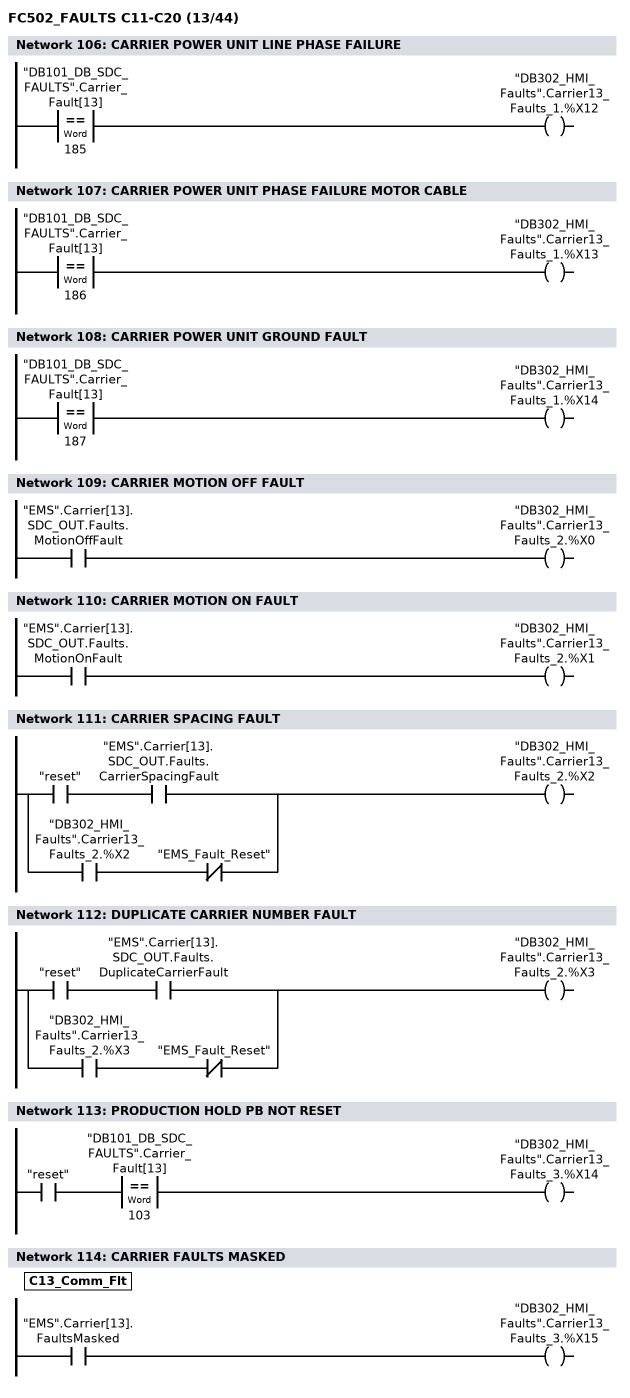
   RUNG wire#powerrail
      { S7_Templates := "SrcType := Word" } EQ_Contact(in1 := "DB101_DB_SDC_FAULTS".Carrier_Fault[13], in2 := 185)
      Coil( "DB302_HMI_Faults".Carrier13_Faults_1.%X12 )
   END_RUNG
   // the same network as SCL:
   "DB302_HMI_Faults".Carrier13_Faults_1.%X12 := "DB101_DB_SDC_FAULTS".Carrier_Fault[13] = 185;
END_REGION

REGION Network 107: CARRIER POWER UNIT PHASE FAILURE MOTOR CABLE
   RUNG wire#powerrail
      { S7_Templates := "SrcType := Word" } EQ_Contact(in1 := "DB101_DB_SDC_FAULTS".Carrier_Fault[13], in2 := 186)
      Coil( "DB302_HMI_Faults".Carrier13_Faults_1.%X13 )
   END_RUNG
   // the same network as SCL:
   "DB302_HMI_Faults".Carrier13_Faults_1.%X13 := "DB101_DB_SDC_FAULTS".Carrier_Fault[13] = 186;
END_REGION

REGION Network 108: CARRIER POWER UNIT GROUND FAULT
   RUNG wire#powerrail
      { S7_Templates := "SrcType := Word" } EQ_Contact(in1 := "DB101_DB_SDC_FAULTS".Carrier_Fault[13], in2 := 187)
      Coil( "DB302_HMI_Faults".Carrier13_Faults_1.%X14 )
   END_RUNG
   // the same network as SCL:
   "DB302_HMI_Faults".Carrier13_Faults_1.%X14 := "DB101_DB_SDC_FAULTS".Carrier_Fault[13] = 187;
END_REGION

REGION Network 109: CARRIER MOTION OFF FAULT
   RUNG wire#powerrail
      Contact( "EMS".Carrier[13].SDC_OUT.Faults.MotionOffFault )
      Coil( "DB302_HMI_Faults".Carrier13_Faults_2.%X0 )
   END_RUNG
   // the same network as SCL:
   "DB302_HMI_Faults".Carrier13_Faults_2.%X0 := "EMS".Carrier[13].SDC_OUT.Faults.MotionOffFault;
END_REGION

REGION Network 110: CARRIER MOTION ON FAULT
   RUNG wire#powerrail
      Contact( "EMS".Carrier[13].SDC_OUT.Faults.MotionOnFault )
      Coil( "DB302_HMI_Faults".Carrier13_Faults_2.%X1 )
   END_RUNG
   // the same network as SCL:
   "DB302_HMI_Faults".Carrier13_Faults_2.%X1 := "EMS".Carrier[13].SDC_OUT.Faults.MotionOnFault;
END_REGION

REGION Network 111: CARRIER SPACING FAULT
   RUNG wire#powerrail
      Contact( "reset" )
      Contact( "EMS".Carrier[13].SDC_OUT.Faults.CarrierSpacingFault )
      wire#w1
      Coil( "DB302_HMI_Faults".Carrier13_Faults_2.%X2 )
   END_RUNG
   RUNG wire#powerrail
      Contact( "DB302_HMI_Faults".Carrier13_Faults_2.%X2 )
      I_Contact( "EMS_Fault_Reset" )
   END_RUNG wire#w1
   // the same network as SCL:
   "DB302_HMI_Faults".Carrier13_Faults_2.%X2 := ("reset" AND "EMS".Carrier[13].SDC_OUT.Faults.CarrierSpacingFault) OR ("DB302_HMI_Faults".Carrier13_Faults_2.%X2 AND NOT "EMS_Fault_Reset");
END_REGION

REGION Network 112: DUPLICATE CARRIER NUMBER FAULT
   RUNG wire#powerrail
      Contact( "reset" )
      Contact( "EMS".Carrier[13].SDC_OUT.Faults.DuplicateCarrierFault )
      wire#w1
      Coil( "DB302_HMI_Faults".Carrier13_Faults_2.%X3 )
   END_RUNG
   RUNG wire#powerrail
      Contact( "DB302_HMI_Faults".Carrier13_Faults_2.%X3 )
      I_Contact( "EMS_Fault_Reset" )
   END_RUNG wire#w1
   // the same network as SCL:
   "DB302_HMI_Faults".Carrier13_Faults_2.%X3 := ("reset" AND "EMS".Carrier[13].SDC_OUT.Faults.DuplicateCarrierFault) OR ("DB302_HMI_Faults".Carrier13_Faults_2.%X3 AND NOT "EMS_Fault_Reset");
END_REGION

REGION Network 113: PRODUCTION HOLD PB NOT RESET
   RUNG wire#powerrail
      Contact( "reset" )
      { S7_Templates := "SrcType := Word" } EQ_Contact(in1 := "DB101_DB_SDC_FAULTS".Carrier_Fault[13], in2 := 103)
      Coil( "DB302_HMI_Faults".Carrier13_Faults_3.%X14 )
   END_RUNG
   // the same network as SCL:
   "DB302_HMI_Faults".Carrier13_Faults_3.%X14 := "reset" AND ("DB101_DB_SDC_FAULTS".Carrier_Fault[13] = 103);
END_REGION

REGION Network 114: CARRIER FAULTS MASKED
   Label( C13_Comm_Flt )
   RUNG wire#powerrail
      Contact( "EMS".Carrier[13].FaultsMasked )
      Coil( "DB302_HMI_Faults".Carrier13_Faults_3.%X15 )
   END_RUNG
   // the same network as SCL:
   C13_Comm_Flt:
   "DB302_HMI_Faults".Carrier13_Faults_3.%X15 := "EMS".Carrier[13].FaultsMasked;
END_REGION

REGION Network 115: CARRIER 14 FAULTS
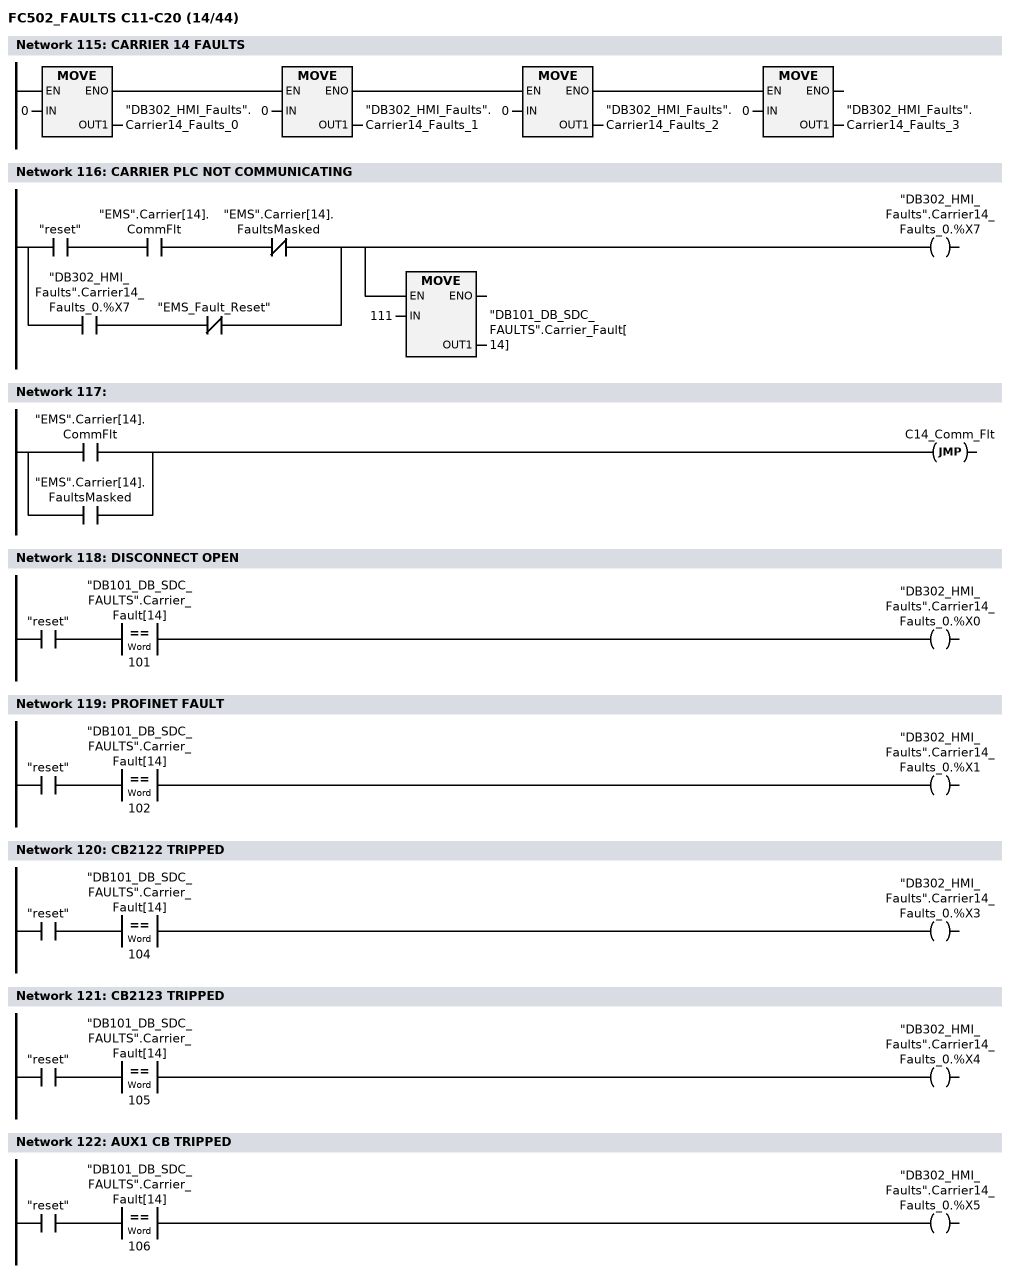
   RUNG wire#powerrail
      Move(in := 0, out1 => "DB302_HMI_Faults".Carrier14_Faults_0)
      Move(in := 0, out1 => "DB302_HMI_Faults".Carrier14_Faults_1)
      Move(in := 0, out1 => "DB302_HMI_Faults".Carrier14_Faults_2)
      Move(in := 0, out1 => "DB302_HMI_Faults".Carrier14_Faults_3)
   END_RUNG
   // the same network as SCL:
   "DB302_HMI_Faults".Carrier14_Faults_0 := 0;
   "DB302_HMI_Faults".Carrier14_Faults_1 := 0;
   "DB302_HMI_Faults".Carrier14_Faults_2 := 0;
   "DB302_HMI_Faults".Carrier14_Faults_3 := 0;
END_REGION

REGION Network 116: CARRIER PLC NOT COMMUNICATING
   RUNG wire#powerrail
      Contact( "reset" )
      Contact( "EMS".Carrier[14].CommFlt )
      I_Contact( "EMS".Carrier[14].FaultsMasked )
      wire#w1
      Coil( "DB302_HMI_Faults".Carrier14_Faults_0.%X7 )
   END_RUNG
   RUNG wire#powerrail
      Contact( "DB302_HMI_Faults".Carrier14_Faults_0.%X7 )
      I_Contact( "EMS_Fault_Reset" )
   END_RUNG wire#w1
   RUNG wire#w1
      Move(in := 111, out1 => "DB101_DB_SDC_FAULTS".Carrier_Fault[14])
   END_RUNG
   // the same network as SCL:
   "DB302_HMI_Faults".Carrier14_Faults_0.%X7 := ("reset" AND "EMS".Carrier[14].CommFlt AND NOT "EMS".Carrier[14].FaultsMasked) OR ("DB302_HMI_Faults".Carrier14_Faults_0.%X7 AND NOT "EMS_Fault_Reset");
   IF "DB302_HMI_Faults".Carrier14_Faults_0.%X7 THEN "DB101_DB_SDC_FAULTS".Carrier_Fault[14] := 111; END_IF;
END_REGION

REGION Network 117
   RUNG wire#powerrail
      Contact( "EMS".Carrier[14].CommFlt )
      wire#w1
      JumpCoil( C14_Comm_Flt )
   END_RUNG
   RUNG wire#powerrail
      Contact( "EMS".Carrier[14].FaultsMasked )
   END_RUNG wire#w1
   // the same network as SCL:
   IF "EMS".Carrier[14].CommFlt OR "EMS".Carrier[14].FaultsMasked THEN GOTO C14_Comm_Flt; END_IF;
END_REGION

REGION Network 118: DISCONNECT OPEN
   RUNG wire#powerrail
      Contact( "reset" )
      { S7_Templates := "SrcType := Word" } EQ_Contact(in1 := "DB101_DB_SDC_FAULTS".Carrier_Fault[14], in2 := 101)
      Coil( "DB302_HMI_Faults".Carrier14_Faults_0.%X0 )
   END_RUNG
   // the same network as SCL:
   "DB302_HMI_Faults".Carrier14_Faults_0.%X0 := "reset" AND ("DB101_DB_SDC_FAULTS".Carrier_Fault[14] = 101);
END_REGION

REGION Network 119: PROFINET FAULT
   RUNG wire#powerrail
      Contact( "reset" )
      { S7_Templates := "SrcType := Word" } EQ_Contact(in1 := "DB101_DB_SDC_FAULTS".Carrier_Fault[14], in2 := 102)
      Coil( "DB302_HMI_Faults".Carrier14_Faults_0.%X1 )
   END_RUNG
   // the same network as SCL:
   "DB302_HMI_Faults".Carrier14_Faults_0.%X1 := "reset" AND ("DB101_DB_SDC_FAULTS".Carrier_Fault[14] = 102);
END_REGION

REGION Network 120: CB2122 TRIPPED
   RUNG wire#powerrail
      Contact( "reset" )
      { S7_Templates := "SrcType := Word" } EQ_Contact(in1 := "DB101_DB_SDC_FAULTS".Carrier_Fault[14], in2 := 104)
      Coil( "DB302_HMI_Faults".Carrier14_Faults_0.%X3 )
   END_RUNG
   // the same network as SCL:
   "DB302_HMI_Faults".Carrier14_Faults_0.%X3 := "reset" AND ("DB101_DB_SDC_FAULTS".Carrier_Fault[14] = 104);
END_REGION

REGION Network 121: CB2123 TRIPPED
   RUNG wire#powerrail
      Contact( "reset" )
      { S7_Templates := "SrcType := Word" } EQ_Contact(in1 := "DB101_DB_SDC_FAULTS".Carrier_Fault[14], in2 := 105)
      Coil( "DB302_HMI_Faults".Carrier14_Faults_0.%X4 )
   END_RUNG
   // the same network as SCL:
   "DB302_HMI_Faults".Carrier14_Faults_0.%X4 := "reset" AND ("DB101_DB_SDC_FAULTS".Carrier_Fault[14] = 105);
END_REGION

REGION Network 122: AUX1 CB TRIPPED
   RUNG wire#powerrail
      Contact( "reset" )
      { S7_Templates := "SrcType := Word" } EQ_Contact(in1 := "DB101_DB_SDC_FAULTS".Carrier_Fault[14], in2 := 106)
      Coil( "DB302_HMI_Faults".Carrier14_Faults_0.%X5 )
   END_RUNG
   // the same network as SCL:
   "DB302_HMI_Faults".Carrier14_Faults_0.%X5 := "reset" AND ("DB101_DB_SDC_FAULTS".Carrier_Fault[14] = 106);
END_REGION

REGION Network 123: AUX2 CB TRIPPED
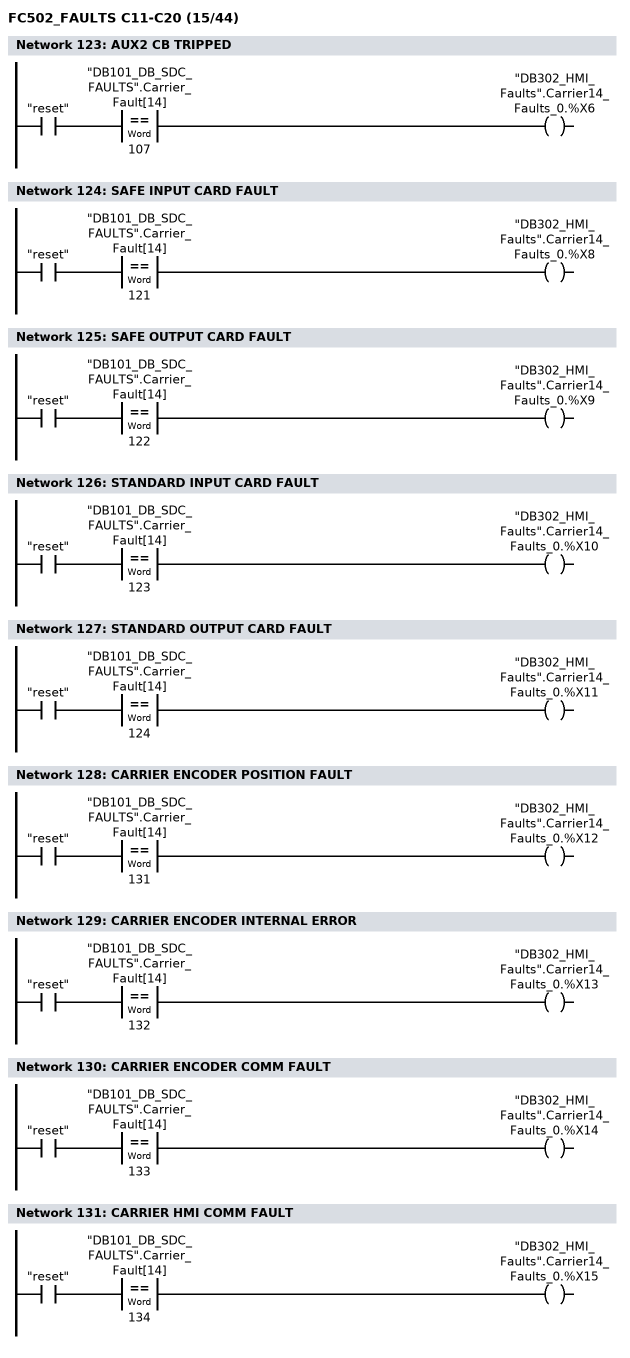
   RUNG wire#powerrail
      Contact( "reset" )
      { S7_Templates := "SrcType := Word" } EQ_Contact(in1 := "DB101_DB_SDC_FAULTS".Carrier_Fault[14], in2 := 107)
      Coil( "DB302_HMI_Faults".Carrier14_Faults_0.%X6 )
   END_RUNG
   // the same network as SCL:
   "DB302_HMI_Faults".Carrier14_Faults_0.%X6 := "reset" AND ("DB101_DB_SDC_FAULTS".Carrier_Fault[14] = 107);
END_REGION

REGION Network 124: SAFE INPUT CARD FAULT
   RUNG wire#powerrail
      Contact( "reset" )
      { S7_Templates := "SrcType := Word" } EQ_Contact(in1 := "DB101_DB_SDC_FAULTS".Carrier_Fault[14], in2 := 121)
      Coil( "DB302_HMI_Faults".Carrier14_Faults_0.%X8 )
   END_RUNG
   // the same network as SCL:
   "DB302_HMI_Faults".Carrier14_Faults_0.%X8 := "reset" AND ("DB101_DB_SDC_FAULTS".Carrier_Fault[14] = 121);
END_REGION

REGION Network 125: SAFE OUTPUT CARD FAULT
   RUNG wire#powerrail
      Contact( "reset" )
      { S7_Templates := "SrcType := Word" } EQ_Contact(in1 := "DB101_DB_SDC_FAULTS".Carrier_Fault[14], in2 := 122)
      Coil( "DB302_HMI_Faults".Carrier14_Faults_0.%X9 )
   END_RUNG
   // the same network as SCL:
   "DB302_HMI_Faults".Carrier14_Faults_0.%X9 := "reset" AND ("DB101_DB_SDC_FAULTS".Carrier_Fault[14] = 122);
END_REGION

REGION Network 126: STANDARD INPUT CARD FAULT
   RUNG wire#powerrail
      Contact( "reset" )
      { S7_Templates := "SrcType := Word" } EQ_Contact(in1 := "DB101_DB_SDC_FAULTS".Carrier_Fault[14], in2 := 123)
      Coil( "DB302_HMI_Faults".Carrier14_Faults_0.%X10 )
   END_RUNG
   // the same network as SCL:
   "DB302_HMI_Faults".Carrier14_Faults_0.%X10 := "reset" AND ("DB101_DB_SDC_FAULTS".Carrier_Fault[14] = 123);
END_REGION

REGION Network 127: STANDARD OUTPUT CARD FAULT
   RUNG wire#powerrail
      Contact( "reset" )
      { S7_Templates := "SrcType := Word" } EQ_Contact(in1 := "DB101_DB_SDC_FAULTS".Carrier_Fault[14], in2 := 124)
      Coil( "DB302_HMI_Faults".Carrier14_Faults_0.%X11 )
   END_RUNG
   // the same network as SCL:
   "DB302_HMI_Faults".Carrier14_Faults_0.%X11 := "reset" AND ("DB101_DB_SDC_FAULTS".Carrier_Fault[14] = 124);
END_REGION

REGION Network 128: CARRIER ENCODER POSITION FAULT
   RUNG wire#powerrail
      Contact( "reset" )
      { S7_Templates := "SrcType := Word" } EQ_Contact(in1 := "DB101_DB_SDC_FAULTS".Carrier_Fault[14], in2 := 131)
      Coil( "DB302_HMI_Faults".Carrier14_Faults_0.%X12 )
   END_RUNG
   // the same network as SCL:
   "DB302_HMI_Faults".Carrier14_Faults_0.%X12 := "reset" AND ("DB101_DB_SDC_FAULTS".Carrier_Fault[14] = 131);
END_REGION

REGION Network 129: CARRIER ENCODER INTERNAL ERROR
   RUNG wire#powerrail
      Contact( "reset" )
      { S7_Templates := "SrcType := Word" } EQ_Contact(in1 := "DB101_DB_SDC_FAULTS".Carrier_Fault[14], in2 := 132)
      Coil( "DB302_HMI_Faults".Carrier14_Faults_0.%X13 )
   END_RUNG
   // the same network as SCL:
   "DB302_HMI_Faults".Carrier14_Faults_0.%X13 := "reset" AND ("DB101_DB_SDC_FAULTS".Carrier_Fault[14] = 132);
END_REGION

REGION Network 130: CARRIER ENCODER COMM FAULT
   RUNG wire#powerrail
      Contact( "reset" )
      { S7_Templates := "SrcType := Word" } EQ_Contact(in1 := "DB101_DB_SDC_FAULTS".Carrier_Fault[14], in2 := 133)
      Coil( "DB302_HMI_Faults".Carrier14_Faults_0.%X14 )
   END_RUNG
   // the same network as SCL:
   "DB302_HMI_Faults".Carrier14_Faults_0.%X14 := "reset" AND ("DB101_DB_SDC_FAULTS".Carrier_Fault[14] = 133);
END_REGION

REGION Network 131: CARRIER HMI COMM FAULT
   RUNG wire#powerrail
      Contact( "reset" )
      { S7_Templates := "SrcType := Word" } EQ_Contact(in1 := "DB101_DB_SDC_FAULTS".Carrier_Fault[14], in2 := 134)
      Coil( "DB302_HMI_Faults".Carrier14_Faults_0.%X15 )
   END_RUNG
   // the same network as SCL:
   "DB302_HMI_Faults".Carrier14_Faults_0.%X15 := "reset" AND ("DB101_DB_SDC_FAULTS".Carrier_Fault[14] = 134);
END_REGION

REGION Network 132: CARRIER CRASH DETECTION FAULT
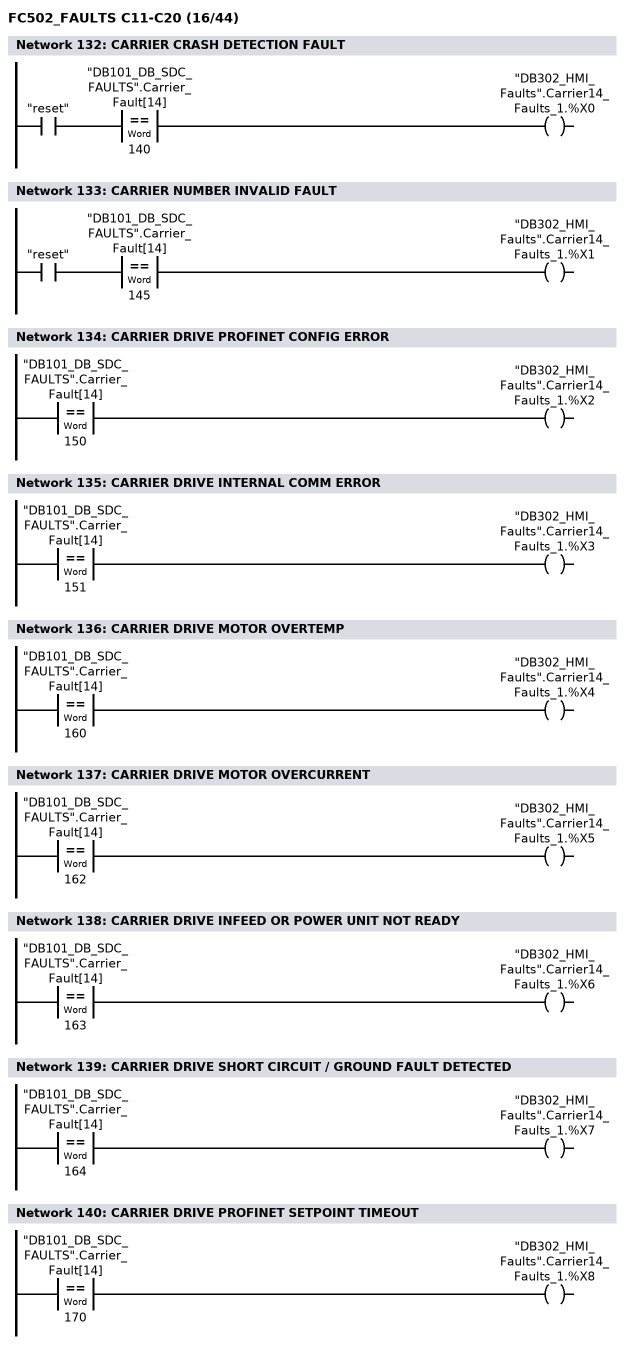
   RUNG wire#powerrail
      Contact( "reset" )
      { S7_Templates := "SrcType := Word" } EQ_Contact(in1 := "DB101_DB_SDC_FAULTS".Carrier_Fault[14], in2 := 140)
      Coil( "DB302_HMI_Faults".Carrier14_Faults_1.%X0 )
   END_RUNG
   // the same network as SCL:
   "DB302_HMI_Faults".Carrier14_Faults_1.%X0 := "reset" AND ("DB101_DB_SDC_FAULTS".Carrier_Fault[14] = 140);
END_REGION

REGION Network 133: CARRIER NUMBER INVALID FAULT
   RUNG wire#powerrail
      Contact( "reset" )
      { S7_Templates := "SrcType := Word" } EQ_Contact(in1 := "DB101_DB_SDC_FAULTS".Carrier_Fault[14], in2 := 145)
      Coil( "DB302_HMI_Faults".Carrier14_Faults_1.%X1 )
   END_RUNG
   // the same network as SCL:
   "DB302_HMI_Faults".Carrier14_Faults_1.%X1 := "reset" AND ("DB101_DB_SDC_FAULTS".Carrier_Fault[14] = 145);
END_REGION

REGION Network 134: CARRIER DRIVE PROFINET CONFIG ERROR
   RUNG wire#powerrail
      { S7_Templates := "SrcType := Word" } EQ_Contact(in1 := "DB101_DB_SDC_FAULTS".Carrier_Fault[14], in2 := 150)
      Coil( "DB302_HMI_Faults".Carrier14_Faults_1.%X2 )
   END_RUNG
   // the same network as SCL:
   "DB302_HMI_Faults".Carrier14_Faults_1.%X2 := "DB101_DB_SDC_FAULTS".Carrier_Fault[14] = 150;
END_REGION

REGION Network 135: CARRIER DRIVE INTERNAL COMM ERROR
   RUNG wire#powerrail
      { S7_Templates := "SrcType := Word" } EQ_Contact(in1 := "DB101_DB_SDC_FAULTS".Carrier_Fault[14], in2 := 151)
      Coil( "DB302_HMI_Faults".Carrier14_Faults_1.%X3 )
   END_RUNG
   // the same network as SCL:
   "DB302_HMI_Faults".Carrier14_Faults_1.%X3 := "DB101_DB_SDC_FAULTS".Carrier_Fault[14] = 151;
END_REGION

REGION Network 136: CARRIER DRIVE MOTOR OVERTEMP
   RUNG wire#powerrail
      { S7_Templates := "SrcType := Word" } EQ_Contact(in1 := "DB101_DB_SDC_FAULTS".Carrier_Fault[14], in2 := 160)
      Coil( "DB302_HMI_Faults".Carrier14_Faults_1.%X4 )
   END_RUNG
   // the same network as SCL:
   "DB302_HMI_Faults".Carrier14_Faults_1.%X4 := "DB101_DB_SDC_FAULTS".Carrier_Fault[14] = 160;
END_REGION

REGION Network 137: CARRIER DRIVE MOTOR OVERCURRENT
   RUNG wire#powerrail
      { S7_Templates := "SrcType := Word" } EQ_Contact(in1 := "DB101_DB_SDC_FAULTS".Carrier_Fault[14], in2 := 162)
      Coil( "DB302_HMI_Faults".Carrier14_Faults_1.%X5 )
   END_RUNG
   // the same network as SCL:
   "DB302_HMI_Faults".Carrier14_Faults_1.%X5 := "DB101_DB_SDC_FAULTS".Carrier_Fault[14] = 162;
END_REGION

REGION Network 138: CARRIER DRIVE INFEED OR POWER UNIT NOT READY
   RUNG wire#powerrail
      { S7_Templates := "SrcType := Word" } EQ_Contact(in1 := "DB101_DB_SDC_FAULTS".Carrier_Fault[14], in2 := 163)
      Coil( "DB302_HMI_Faults".Carrier14_Faults_1.%X6 )
   END_RUNG
   // the same network as SCL:
   "DB302_HMI_Faults".Carrier14_Faults_1.%X6 := "DB101_DB_SDC_FAULTS".Carrier_Fault[14] = 163;
END_REGION

REGION Network 139: CARRIER DRIVE SHORT CIRCUIT / GROUND FAULT DETECTED
   RUNG wire#powerrail
      { S7_Templates := "SrcType := Word" } EQ_Contact(in1 := "DB101_DB_SDC_FAULTS".Carrier_Fault[14], in2 := 164)
      Coil( "DB302_HMI_Faults".Carrier14_Faults_1.%X7 )
   END_RUNG
   // the same network as SCL:
   "DB302_HMI_Faults".Carrier14_Faults_1.%X7 := "DB101_DB_SDC_FAULTS".Carrier_Fault[14] = 164;
END_REGION

REGION Network 140: CARRIER DRIVE PROFINET SETPOINT TIMEOUT
   RUNG wire#powerrail
      { S7_Templates := "SrcType := Word" } EQ_Contact(in1 := "DB101_DB_SDC_FAULTS".Carrier_Fault[14], in2 := 170)
      Coil( "DB302_HMI_Faults".Carrier14_Faults_1.%X8 )
   END_RUNG
   // the same network as SCL:
   "DB302_HMI_Faults".Carrier14_Faults_1.%X8 := "DB101_DB_SDC_FAULTS".Carrier_Fault[14] = 170;
END_REGION

REGION Network 141: CARRIER POWER UNIT OVERCURRENT
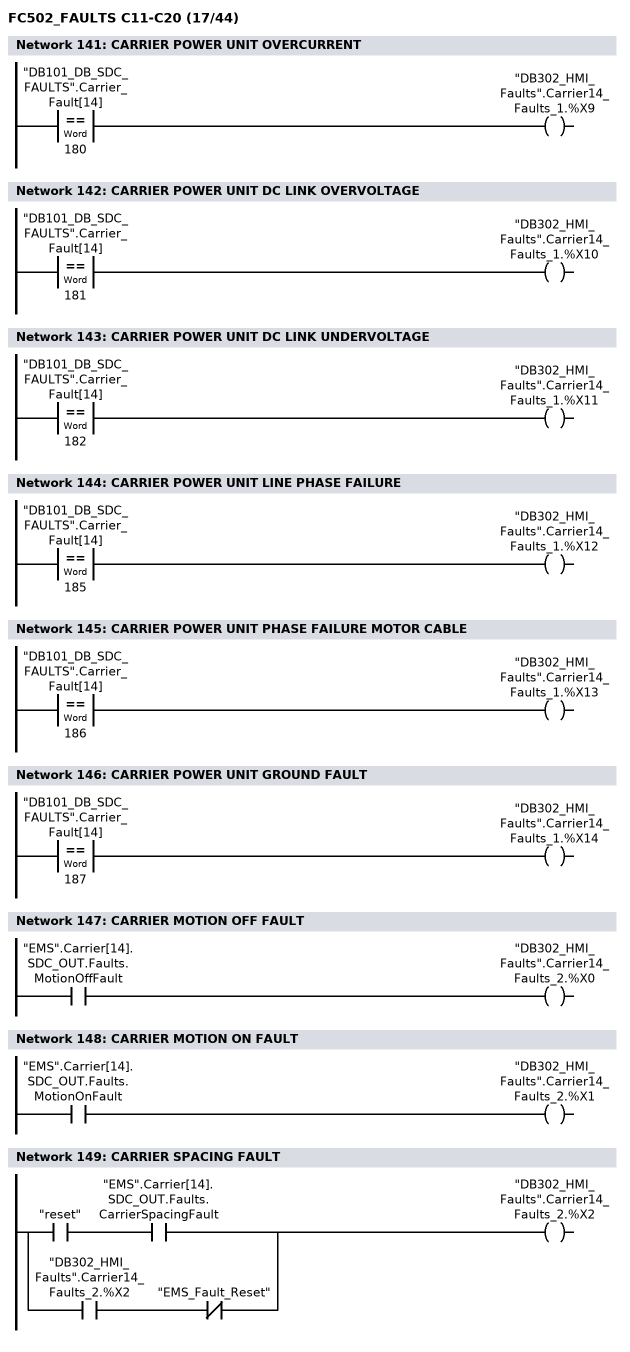
   RUNG wire#powerrail
      { S7_Templates := "SrcType := Word" } EQ_Contact(in1 := "DB101_DB_SDC_FAULTS".Carrier_Fault[14], in2 := 180)
      Coil( "DB302_HMI_Faults".Carrier14_Faults_1.%X9 )
   END_RUNG
   // the same network as SCL:
   "DB302_HMI_Faults".Carrier14_Faults_1.%X9 := "DB101_DB_SDC_FAULTS".Carrier_Fault[14] = 180;
END_REGION

REGION Network 142: CARRIER POWER UNIT DC LINK OVERVOLTAGE
   RUNG wire#powerrail
      { S7_Templates := "SrcType := Word" } EQ_Contact(in1 := "DB101_DB_SDC_FAULTS".Carrier_Fault[14], in2 := 181)
      Coil( "DB302_HMI_Faults".Carrier14_Faults_1.%X10 )
   END_RUNG
   // the same network as SCL:
   "DB302_HMI_Faults".Carrier14_Faults_1.%X10 := "DB101_DB_SDC_FAULTS".Carrier_Fault[14] = 181;
END_REGION

REGION Network 143: CARRIER POWER UNIT DC LINK UNDERVOLTAGE
   RUNG wire#powerrail
      { S7_Templates := "SrcType := Word" } EQ_Contact(in1 := "DB101_DB_SDC_FAULTS".Carrier_Fault[14], in2 := 182)
      Coil( "DB302_HMI_Faults".Carrier14_Faults_1.%X11 )
   END_RUNG
   // the same network as SCL:
   "DB302_HMI_Faults".Carrier14_Faults_1.%X11 := "DB101_DB_SDC_FAULTS".Carrier_Fault[14] = 182;
END_REGION

REGION Network 144: CARRIER POWER UNIT LINE PHASE FAILURE
   RUNG wire#powerrail
      { S7_Templates := "SrcType := Word" } EQ_Contact(in1 := "DB101_DB_SDC_FAULTS".Carrier_Fault[14], in2 := 185)
      Coil( "DB302_HMI_Faults".Carrier14_Faults_1.%X12 )
   END_RUNG
   // the same network as SCL:
   "DB302_HMI_Faults".Carrier14_Faults_1.%X12 := "DB101_DB_SDC_FAULTS".Carrier_Fault[14] = 185;
END_REGION

REGION Network 145: CARRIER POWER UNIT PHASE FAILURE MOTOR CABLE
   RUNG wire#powerrail
      { S7_Templates := "SrcType := Word" } EQ_Contact(in1 := "DB101_DB_SDC_FAULTS".Carrier_Fault[14], in2 := 186)
      Coil( "DB302_HMI_Faults".Carrier14_Faults_1.%X13 )
   END_RUNG
   // the same network as SCL:
   "DB302_HMI_Faults".Carrier14_Faults_1.%X13 := "DB101_DB_SDC_FAULTS".Carrier_Fault[14] = 186;
END_REGION

REGION Network 146: CARRIER POWER UNIT GROUND FAULT
   RUNG wire#powerrail
      { S7_Templates := "SrcType := Word" } EQ_Contact(in1 := "DB101_DB_SDC_FAULTS".Carrier_Fault[14], in2 := 187)
      Coil( "DB302_HMI_Faults".Carrier14_Faults_1.%X14 )
   END_RUNG
   // the same network as SCL:
   "DB302_HMI_Faults".Carrier14_Faults_1.%X14 := "DB101_DB_SDC_FAULTS".Carrier_Fault[14] = 187;
END_REGION

REGION Network 147: CARRIER MOTION OFF FAULT
   RUNG wire#powerrail
      Contact( "EMS".Carrier[14].SDC_OUT.Faults.MotionOffFault )
      Coil( "DB302_HMI_Faults".Carrier14_Faults_2.%X0 )
   END_RUNG
   // the same network as SCL:
   "DB302_HMI_Faults".Carrier14_Faults_2.%X0 := "EMS".Carrier[14].SDC_OUT.Faults.MotionOffFault;
END_REGION

REGION Network 148: CARRIER MOTION ON FAULT
   RUNG wire#powerrail
      Contact( "EMS".Carrier[14].SDC_OUT.Faults.MotionOnFault )
      Coil( "DB302_HMI_Faults".Carrier14_Faults_2.%X1 )
   END_RUNG
   // the same network as SCL:
   "DB302_HMI_Faults".Carrier14_Faults_2.%X1 := "EMS".Carrier[14].SDC_OUT.Faults.MotionOnFault;
END_REGION

REGION Network 149: CARRIER SPACING FAULT
   RUNG wire#powerrail
      Contact( "reset" )
      Contact( "EMS".Carrier[14].SDC_OUT.Faults.CarrierSpacingFault )
      wire#w1
      Coil( "DB302_HMI_Faults".Carrier14_Faults_2.%X2 )
   END_RUNG
   RUNG wire#powerrail
      Contact( "DB302_HMI_Faults".Carrier14_Faults_2.%X2 )
      I_Contact( "EMS_Fault_Reset" )
   END_RUNG wire#w1
   // the same network as SCL:
   "DB302_HMI_Faults".Carrier14_Faults_2.%X2 := ("reset" AND "EMS".Carrier[14].SDC_OUT.Faults.CarrierSpacingFault) OR ("DB302_HMI_Faults".Carrier14_Faults_2.%X2 AND NOT "EMS_Fault_Reset");
END_REGION

REGION Network 150: DUPLICATE CARRIER NUMBER FAULT
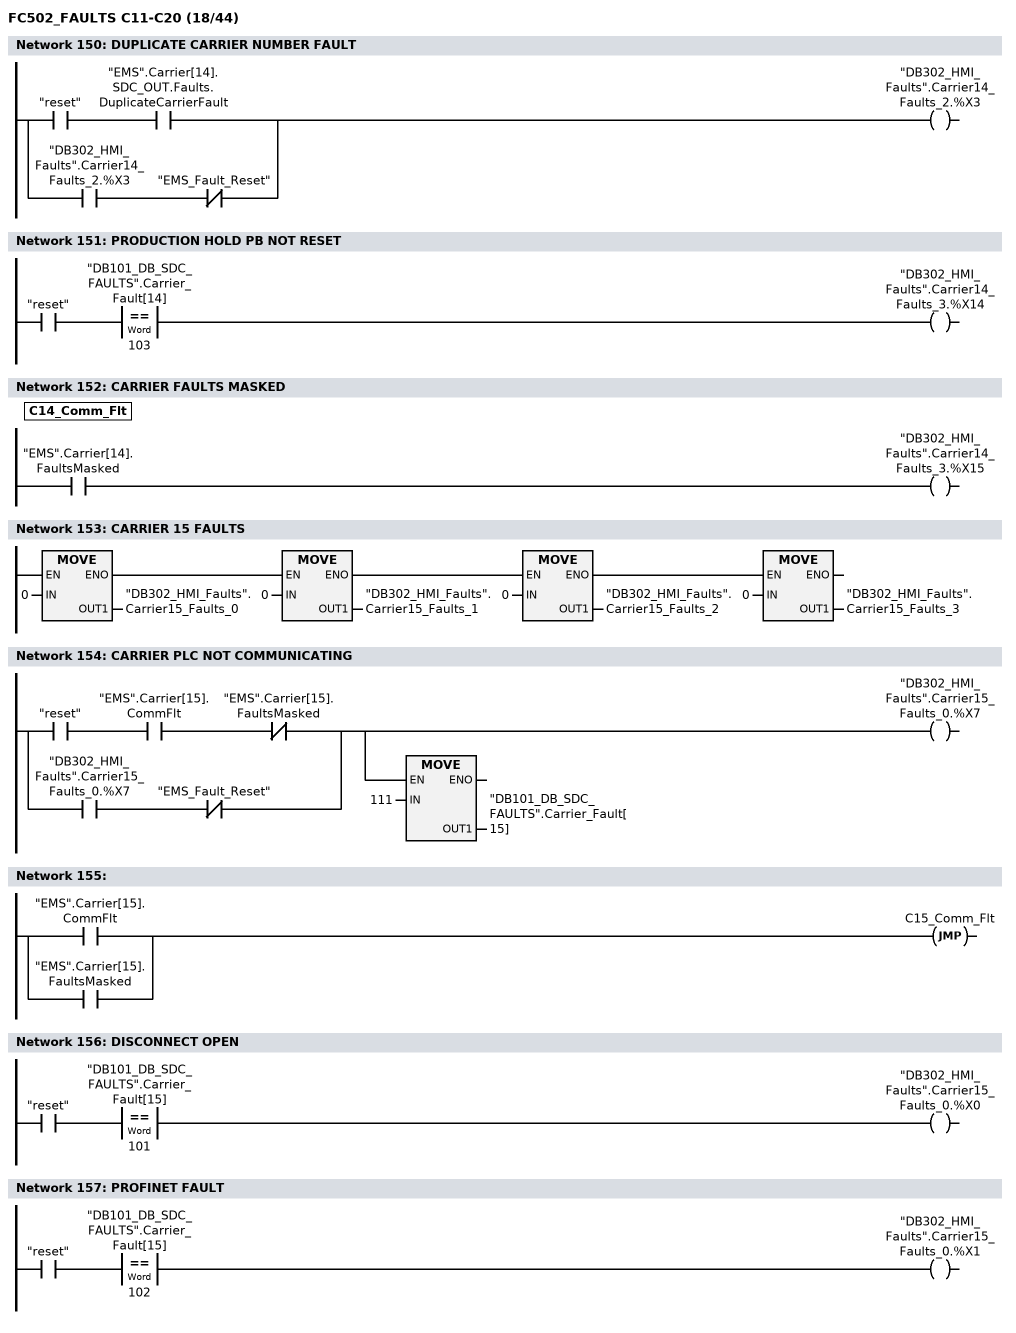
   RUNG wire#powerrail
      Contact( "reset" )
      Contact( "EMS".Carrier[14].SDC_OUT.Faults.DuplicateCarrierFault )
      wire#w1
      Coil( "DB302_HMI_Faults".Carrier14_Faults_2.%X3 )
   END_RUNG
   RUNG wire#powerrail
      Contact( "DB302_HMI_Faults".Carrier14_Faults_2.%X3 )
      I_Contact( "EMS_Fault_Reset" )
   END_RUNG wire#w1
   // the same network as SCL:
   "DB302_HMI_Faults".Carrier14_Faults_2.%X3 := ("reset" AND "EMS".Carrier[14].SDC_OUT.Faults.DuplicateCarrierFault) OR ("DB302_HMI_Faults".Carrier14_Faults_2.%X3 AND NOT "EMS_Fault_Reset");
END_REGION

REGION Network 151: PRODUCTION HOLD PB NOT RESET
   RUNG wire#powerrail
      Contact( "reset" )
      { S7_Templates := "SrcType := Word" } EQ_Contact(in1 := "DB101_DB_SDC_FAULTS".Carrier_Fault[14], in2 := 103)
      Coil( "DB302_HMI_Faults".Carrier14_Faults_3.%X14 )
   END_RUNG
   // the same network as SCL:
   "DB302_HMI_Faults".Carrier14_Faults_3.%X14 := "reset" AND ("DB101_DB_SDC_FAULTS".Carrier_Fault[14] = 103);
END_REGION

REGION Network 152: CARRIER FAULTS MASKED
   Label( C14_Comm_Flt )
   RUNG wire#powerrail
      Contact( "EMS".Carrier[14].FaultsMasked )
      Coil( "DB302_HMI_Faults".Carrier14_Faults_3.%X15 )
   END_RUNG
   // the same network as SCL:
   C14_Comm_Flt:
   "DB302_HMI_Faults".Carrier14_Faults_3.%X15 := "EMS".Carrier[14].FaultsMasked;
END_REGION

REGION Network 153: CARRIER 15 FAULTS
   RUNG wire#powerrail
      Move(in := 0, out1 => "DB302_HMI_Faults".Carrier15_Faults_0)
      Move(in := 0, out1 => "DB302_HMI_Faults".Carrier15_Faults_1)
      Move(in := 0, out1 => "DB302_HMI_Faults".Carrier15_Faults_2)
      Move(in := 0, out1 => "DB302_HMI_Faults".Carrier15_Faults_3)
   END_RUNG
   // the same network as SCL:
   "DB302_HMI_Faults".Carrier15_Faults_0 := 0;
   "DB302_HMI_Faults".Carrier15_Faults_1 := 0;
   "DB302_HMI_Faults".Carrier15_Faults_2 := 0;
   "DB302_HMI_Faults".Carrier15_Faults_3 := 0;
END_REGION

REGION Network 154: CARRIER PLC NOT COMMUNICATING
   RUNG wire#powerrail
      Contact( "reset" )
      Contact( "EMS".Carrier[15].CommFlt )
      I_Contact( "EMS".Carrier[15].FaultsMasked )
      wire#w1
      Coil( "DB302_HMI_Faults".Carrier15_Faults_0.%X7 )
   END_RUNG
   RUNG wire#powerrail
      Contact( "DB302_HMI_Faults".Carrier15_Faults_0.%X7 )
      I_Contact( "EMS_Fault_Reset" )
   END_RUNG wire#w1
   RUNG wire#w1
      Move(in := 111, out1 => "DB101_DB_SDC_FAULTS".Carrier_Fault[15])
   END_RUNG
   // the same network as SCL:
   "DB302_HMI_Faults".Carrier15_Faults_0.%X7 := ("reset" AND "EMS".Carrier[15].CommFlt AND NOT "EMS".Carrier[15].FaultsMasked) OR ("DB302_HMI_Faults".Carrier15_Faults_0.%X7 AND NOT "EMS_Fault_Reset");
   IF "DB302_HMI_Faults".Carrier15_Faults_0.%X7 THEN "DB101_DB_SDC_FAULTS".Carrier_Fault[15] := 111; END_IF;
END_REGION

REGION Network 155
   RUNG wire#powerrail
      Contact( "EMS".Carrier[15].CommFlt )
      wire#w1
      JumpCoil( C15_Comm_Flt )
   END_RUNG
   RUNG wire#powerrail
      Contact( "EMS".Carrier[15].FaultsMasked )
   END_RUNG wire#w1
   // the same network as SCL:
   IF "EMS".Carrier[15].CommFlt OR "EMS".Carrier[15].FaultsMasked THEN GOTO C15_Comm_Flt; END_IF;
END_REGION

REGION Network 156: DISCONNECT OPEN
   RUNG wire#powerrail
      Contact( "reset" )
      { S7_Templates := "SrcType := Word" } EQ_Contact(in1 := "DB101_DB_SDC_FAULTS".Carrier_Fault[15], in2 := 101)
      Coil( "DB302_HMI_Faults".Carrier15_Faults_0.%X0 )
   END_RUNG
   // the same network as SCL:
   "DB302_HMI_Faults".Carrier15_Faults_0.%X0 := "reset" AND ("DB101_DB_SDC_FAULTS".Carrier_Fault[15] = 101);
END_REGION

REGION Network 157: PROFINET FAULT
   RUNG wire#powerrail
      Contact( "reset" )
      { S7_Templates := "SrcType := Word" } EQ_Contact(in1 := "DB101_DB_SDC_FAULTS".Carrier_Fault[15], in2 := 102)
      Coil( "DB302_HMI_Faults".Carrier15_Faults_0.%X1 )
   END_RUNG
   // the same network as SCL:
   "DB302_HMI_Faults".Carrier15_Faults_0.%X1 := "reset" AND ("DB101_DB_SDC_FAULTS".Carrier_Fault[15] = 102);
END_REGION

REGION Network 158: CB2122 TRIPPED
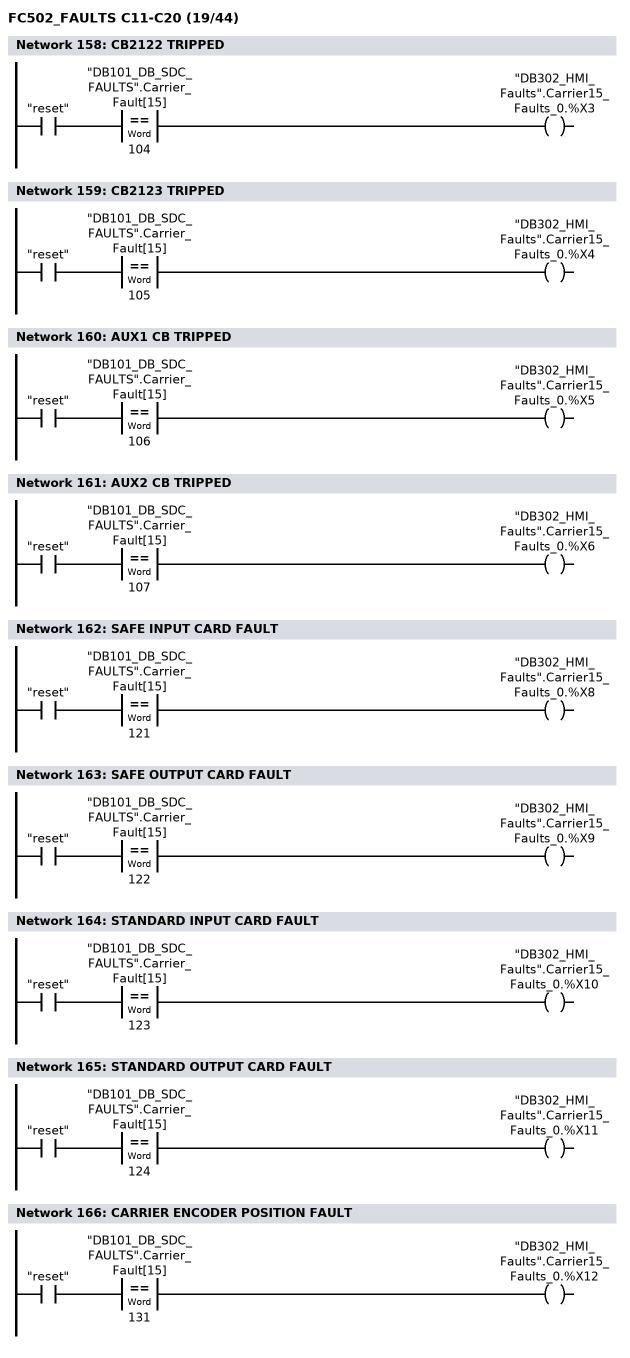
   RUNG wire#powerrail
      Contact( "reset" )
      { S7_Templates := "SrcType := Word" } EQ_Contact(in1 := "DB101_DB_SDC_FAULTS".Carrier_Fault[15], in2 := 104)
      Coil( "DB302_HMI_Faults".Carrier15_Faults_0.%X3 )
   END_RUNG
   // the same network as SCL:
   "DB302_HMI_Faults".Carrier15_Faults_0.%X3 := "reset" AND ("DB101_DB_SDC_FAULTS".Carrier_Fault[15] = 104);
END_REGION

REGION Network 159: CB2123 TRIPPED
   RUNG wire#powerrail
      Contact( "reset" )
      { S7_Templates := "SrcType := Word" } EQ_Contact(in1 := "DB101_DB_SDC_FAULTS".Carrier_Fault[15], in2 := 105)
      Coil( "DB302_HMI_Faults".Carrier15_Faults_0.%X4 )
   END_RUNG
   // the same network as SCL:
   "DB302_HMI_Faults".Carrier15_Faults_0.%X4 := "reset" AND ("DB101_DB_SDC_FAULTS".Carrier_Fault[15] = 105);
END_REGION

REGION Network 160: AUX1 CB TRIPPED
   RUNG wire#powerrail
      Contact( "reset" )
      { S7_Templates := "SrcType := Word" } EQ_Contact(in1 := "DB101_DB_SDC_FAULTS".Carrier_Fault[15], in2 := 106)
      Coil( "DB302_HMI_Faults".Carrier15_Faults_0.%X5 )
   END_RUNG
   // the same network as SCL:
   "DB302_HMI_Faults".Carrier15_Faults_0.%X5 := "reset" AND ("DB101_DB_SDC_FAULTS".Carrier_Fault[15] = 106);
END_REGION

REGION Network 161: AUX2 CB TRIPPED
   RUNG wire#powerrail
      Contact( "reset" )
      { S7_Templates := "SrcType := Word" } EQ_Contact(in1 := "DB101_DB_SDC_FAULTS".Carrier_Fault[15], in2 := 107)
      Coil( "DB302_HMI_Faults".Carrier15_Faults_0.%X6 )
   END_RUNG
   // the same network as SCL:
   "DB302_HMI_Faults".Carrier15_Faults_0.%X6 := "reset" AND ("DB101_DB_SDC_FAULTS".Carrier_Fault[15] = 107);
END_REGION

REGION Network 162: SAFE INPUT CARD FAULT
   RUNG wire#powerrail
      Contact( "reset" )
      { S7_Templates := "SrcType := Word" } EQ_Contact(in1 := "DB101_DB_SDC_FAULTS".Carrier_Fault[15], in2 := 121)
      Coil( "DB302_HMI_Faults".Carrier15_Faults_0.%X8 )
   END_RUNG
   // the same network as SCL:
   "DB302_HMI_Faults".Carrier15_Faults_0.%X8 := "reset" AND ("DB101_DB_SDC_FAULTS".Carrier_Fault[15] = 121);
END_REGION

REGION Network 163: SAFE OUTPUT CARD FAULT
   RUNG wire#powerrail
      Contact( "reset" )
      { S7_Templates := "SrcType := Word" } EQ_Contact(in1 := "DB101_DB_SDC_FAULTS".Carrier_Fault[15], in2 := 122)
      Coil( "DB302_HMI_Faults".Carrier15_Faults_0.%X9 )
   END_RUNG
   // the same network as SCL:
   "DB302_HMI_Faults".Carrier15_Faults_0.%X9 := "reset" AND ("DB101_DB_SDC_FAULTS".Carrier_Fault[15] = 122);
END_REGION

REGION Network 164: STANDARD INPUT CARD FAULT
   RUNG wire#powerrail
      Contact( "reset" )
      { S7_Templates := "SrcType := Word" } EQ_Contact(in1 := "DB101_DB_SDC_FAULTS".Carrier_Fault[15], in2 := 123)
      Coil( "DB302_HMI_Faults".Carrier15_Faults_0.%X10 )
   END_RUNG
   // the same network as SCL:
   "DB302_HMI_Faults".Carrier15_Faults_0.%X10 := "reset" AND ("DB101_DB_SDC_FAULTS".Carrier_Fault[15] = 123);
END_REGION

REGION Network 165: STANDARD OUTPUT CARD FAULT
   RUNG wire#powerrail
      Contact( "reset" )
      { S7_Templates := "SrcType := Word" } EQ_Contact(in1 := "DB101_DB_SDC_FAULTS".Carrier_Fault[15], in2 := 124)
      Coil( "DB302_HMI_Faults".Carrier15_Faults_0.%X11 )
   END_RUNG
   // the same network as SCL:
   "DB302_HMI_Faults".Carrier15_Faults_0.%X11 := "reset" AND ("DB101_DB_SDC_FAULTS".Carrier_Fault[15] = 124);
END_REGION

REGION Network 166: CARRIER ENCODER POSITION FAULT
   RUNG wire#powerrail
      Contact( "reset" )
      { S7_Templates := "SrcType := Word" } EQ_Contact(in1 := "DB101_DB_SDC_FAULTS".Carrier_Fault[15], in2 := 131)
      Coil( "DB302_HMI_Faults".Carrier15_Faults_0.%X12 )
   END_RUNG
   // the same network as SCL:
   "DB302_HMI_Faults".Carrier15_Faults_0.%X12 := "reset" AND ("DB101_DB_SDC_FAULTS".Carrier_Fault[15] = 131);
END_REGION

REGION Network 167: CARRIER ENCODER INTERNAL ERROR
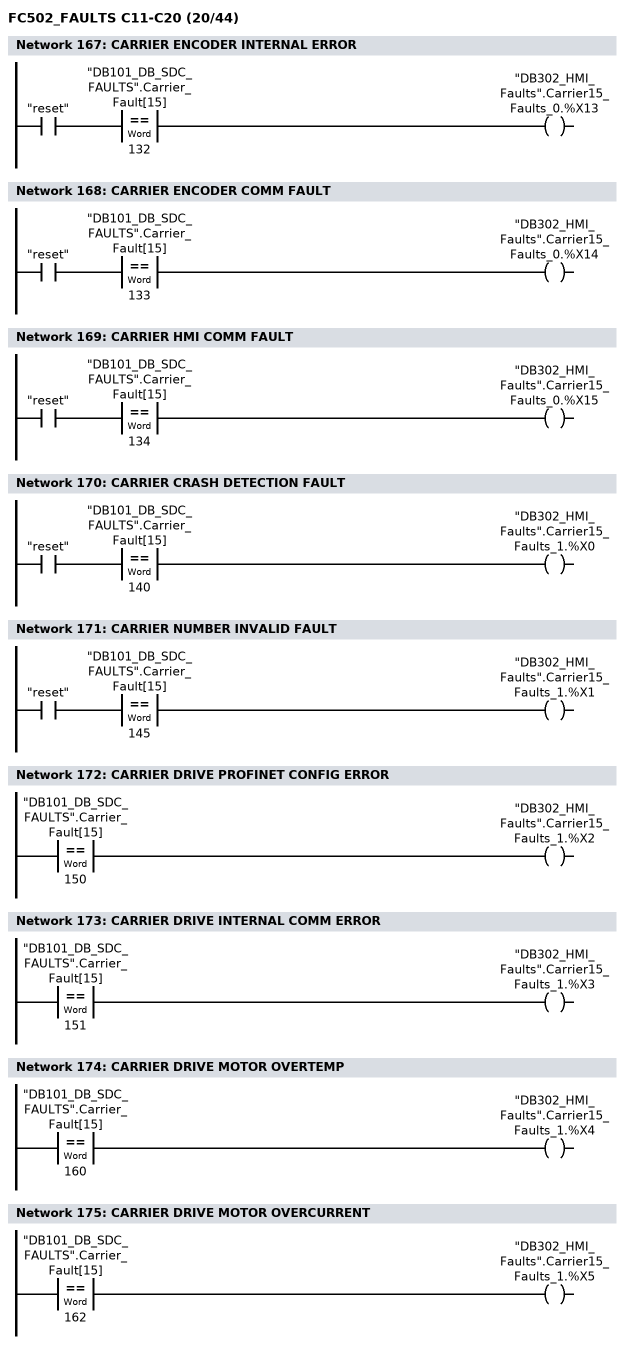
   RUNG wire#powerrail
      Contact( "reset" )
      { S7_Templates := "SrcType := Word" } EQ_Contact(in1 := "DB101_DB_SDC_FAULTS".Carrier_Fault[15], in2 := 132)
      Coil( "DB302_HMI_Faults".Carrier15_Faults_0.%X13 )
   END_RUNG
   // the same network as SCL:
   "DB302_HMI_Faults".Carrier15_Faults_0.%X13 := "reset" AND ("DB101_DB_SDC_FAULTS".Carrier_Fault[15] = 132);
END_REGION

REGION Network 168: CARRIER ENCODER COMM FAULT
   RUNG wire#powerrail
      Contact( "reset" )
      { S7_Templates := "SrcType := Word" } EQ_Contact(in1 := "DB101_DB_SDC_FAULTS".Carrier_Fault[15], in2 := 133)
      Coil( "DB302_HMI_Faults".Carrier15_Faults_0.%X14 )
   END_RUNG
   // the same network as SCL:
   "DB302_HMI_Faults".Carrier15_Faults_0.%X14 := "reset" AND ("DB101_DB_SDC_FAULTS".Carrier_Fault[15] = 133);
END_REGION

REGION Network 169: CARRIER HMI COMM FAULT
   RUNG wire#powerrail
      Contact( "reset" )
      { S7_Templates := "SrcType := Word" } EQ_Contact(in1 := "DB101_DB_SDC_FAULTS".Carrier_Fault[15], in2 := 134)
      Coil( "DB302_HMI_Faults".Carrier15_Faults_0.%X15 )
   END_RUNG
   // the same network as SCL:
   "DB302_HMI_Faults".Carrier15_Faults_0.%X15 := "reset" AND ("DB101_DB_SDC_FAULTS".Carrier_Fault[15] = 134);
END_REGION

REGION Network 170: CARRIER CRASH DETECTION FAULT
   RUNG wire#powerrail
      Contact( "reset" )
      { S7_Templates := "SrcType := Word" } EQ_Contact(in1 := "DB101_DB_SDC_FAULTS".Carrier_Fault[15], in2 := 140)
      Coil( "DB302_HMI_Faults".Carrier15_Faults_1.%X0 )
   END_RUNG
   // the same network as SCL:
   "DB302_HMI_Faults".Carrier15_Faults_1.%X0 := "reset" AND ("DB101_DB_SDC_FAULTS".Carrier_Fault[15] = 140);
END_REGION

REGION Network 171: CARRIER NUMBER INVALID FAULT
   RUNG wire#powerrail
      Contact( "reset" )
      { S7_Templates := "SrcType := Word" } EQ_Contact(in1 := "DB101_DB_SDC_FAULTS".Carrier_Fault[15], in2 := 145)
      Coil( "DB302_HMI_Faults".Carrier15_Faults_1.%X1 )
   END_RUNG
   // the same network as SCL:
   "DB302_HMI_Faults".Carrier15_Faults_1.%X1 := "reset" AND ("DB101_DB_SDC_FAULTS".Carrier_Fault[15] = 145);
END_REGION

REGION Network 172: CARRIER DRIVE PROFINET CONFIG ERROR
   RUNG wire#powerrail
      { S7_Templates := "SrcType := Word" } EQ_Contact(in1 := "DB101_DB_SDC_FAULTS".Carrier_Fault[15], in2 := 150)
      Coil( "DB302_HMI_Faults".Carrier15_Faults_1.%X2 )
   END_RUNG
   // the same network as SCL:
   "DB302_HMI_Faults".Carrier15_Faults_1.%X2 := "DB101_DB_SDC_FAULTS".Carrier_Fault[15] = 150;
END_REGION

REGION Network 173: CARRIER DRIVE INTERNAL COMM ERROR
   RUNG wire#powerrail
      { S7_Templates := "SrcType := Word" } EQ_Contact(in1 := "DB101_DB_SDC_FAULTS".Carrier_Fault[15], in2 := 151)
      Coil( "DB302_HMI_Faults".Carrier15_Faults_1.%X3 )
   END_RUNG
   // the same network as SCL:
   "DB302_HMI_Faults".Carrier15_Faults_1.%X3 := "DB101_DB_SDC_FAULTS".Carrier_Fault[15] = 151;
END_REGION

REGION Network 174: CARRIER DRIVE MOTOR OVERTEMP
   RUNG wire#powerrail
      { S7_Templates := "SrcType := Word" } EQ_Contact(in1 := "DB101_DB_SDC_FAULTS".Carrier_Fault[15], in2 := 160)
      Coil( "DB302_HMI_Faults".Carrier15_Faults_1.%X4 )
   END_RUNG
   // the same network as SCL:
   "DB302_HMI_Faults".Carrier15_Faults_1.%X4 := "DB101_DB_SDC_FAULTS".Carrier_Fault[15] = 160;
END_REGION

REGION Network 175: CARRIER DRIVE MOTOR OVERCURRENT
   RUNG wire#powerrail
      { S7_Templates := "SrcType := Word" } EQ_Contact(in1 := "DB101_DB_SDC_FAULTS".Carrier_Fault[15], in2 := 162)
      Coil( "DB302_HMI_Faults".Carrier15_Faults_1.%X5 )
   END_RUNG
   // the same network as SCL:
   "DB302_HMI_Faults".Carrier15_Faults_1.%X5 := "DB101_DB_SDC_FAULTS".Carrier_Fault[15] = 162;
END_REGION

REGION Network 176: CARRIER DRIVE INFEED OR POWER UNIT NOT READY
